Controller 1 Volume Not Ok Fault FB1[260].20'; 8341 '~S001R03CN.I.Slr1PurgeFlt - Seal Controller 1 Purge Fault FB1[260].21'; 8342 '~S001R03CN.I.Slr1DoserNot Filled - Seal Cntrl 1 Doser Not Filled FB1[260].22'; 8343 '~S001R03CN.I.Slr1No2ClnMxr - Seal Cntrl1 No 2C In Mixer Fault FB1[260].23'; 8344 '~S001R03CN.I.Slr1NzlBroken - Seal Controller 1 Nozzle Broken Fault FB1[260].24'; 8345 '~S001R03CN.I.Slr1NozzleChgReq - Seal Cntrl1 Nozzle Change Reqd FB1[260].25'; 8346 '~S001R03CN.I.Slr1CycleInterrupted - Seal Cntrl1 Cycle Interrupted FB1[260].26'; 8347 '~S001R03CN.I.Stdw1Flt - Stud Weld 1 Weld Fault FB1[260].27'; 8348 '~S001R03CN.I.Stdw1DlyExcdd - Stud Weld 1 Time Delay Exceeded Flt FB1[260].28'; 8349 '~S001R03CN.I.Stdw1Maint Reqd - Stud Weld 1 Maintenance Required FB1[260].29'; 8350 '~S001R03CN.I.Stdw1Reject - Stud Weld 1 art Reject Fault FB1[260].30'; 8351 '~S001R03CN.I.Rvt1Flt - Rivet Controller 1 Fault FB1[260].31'; 8352 '~S001R03CN.I.Rvt1DlyExcdd - Rivet Cntrl 1 Time Delay Exceeded Flt FB1[261].0'; 8353 '~S001R03CN.I.AutoPulledTipByp1 - Auto Pulled Tip Bypass 1 FB1[261].1'; 8354 '~S001R03CN.I.StdWld1EquipmentFlt - Stud Weld 1 Equipment Fault FB1[261].2'; 8355 '~S001R03CN.I.StdWld1BrcktNotPresent - Stud Weld 1 Bracket Not Pres FB1[261].3'; 8356 '~S001R03CN.I.PierceFlt - Pierce Fault FB1[261].4'; 8357 '~S001R03CN.I.NoVisionMeasErr - Vision System Measurement Error FB1[261].5'; 8358 '~S001R03CN.I.VisionSysCalErr - Vision System Calibration Fault FB1[261].6'; 8359 '~S001R03CN.I.VisionSysErr - Vision System Error FB1[261].7'; 8360 '~S001R03CN.I.RackOutOfTolerance - Vision Sys Rack Out Of Tolerance FB1[261].8'; 8361 '~S001R03CN.Ix.TorqFlt - Torque Not Ok FB1[261].9'; 8362 '~S001R03CN.Ix.MwFlt - Mig Weld Controller Fault FB1[261].10'; 8363 '~S001R03CN.Ix.MwWireStuckFlt - Mig Welder Wire Stuck FB1[261].11'; 8364 '~S001R03CN.Ix.MwWldFlt - Mig Welder Bad Bronze Weld Indicator Flt FB1[261].12'; 8365 '~S001R03CN.I.O.TipChngReqd1 - Weld Cntrl 1 Tip Change Required FB1[261].13'; 8366 '~S001R03CN.I.M.NutDetectFlt1 - Nut Welder 1 Nut Detection Fault FB1[261].14'; 8367 '~S001R03CN.I.M.NutProjFlt1 - Nut Welder 1 Weld Not In Tolerance FB1[261].15'; 8368 '~S001R03CN.M.WrongRivetAtNose - Remove Wrong Rivet At Nose FB1[261].16'; 8369 '~S001R03CN.Ix.MwWldLimitErr - Mig Welder CurrentVoltage Out of Tolerance FB1[261].17'; 8370 '~S001R03CN.Ix.MigRdy Mig Welder Not Ready FB1[261].18'; 8371 '~Spare FB1[261].19'; 8372 '~Spare FB1[261].20'; 8373 '~S001R03CN.I.Wc2WldFlt -Weld Controller 2 Weld Fault FB1[261].21'; 8374 '~S001R03CN.I.Wc2Flt - Weld Timer Flt - Depress Man Weld To Continue FB1[261].22'; 8375 '~S001R03CN.I.Wc2SGunFlt - Weld Controller 2 Servo Gun Fault FB1[261].23'; 8376 '~S001R03CN.I.Wc2SGunMtrTempFlt - Cntrl 2 Servo Gun Motor Over Temp FB1[261].24'; 8377 '~S001R03CN.I.Td2MtrFlt - Tip Dress 2 Motor Fault FB1[261].25'; 8378 '~S001R03CN.I.WC2XfmrTempFlt - Weld Cntrl 2 Transformer Over Temp FB1[261].26'; 8379 '~S001R03CN.I.AutoTipChng2Flt - Auto Tip Changer 2 Fault FB1[261].27'; 8380 '~S001R03CN.I.Slr2NotReady - Seal Controller 2 Not Ready FB1[261].28'; 8381 '~S001R03CN.I.Slr2MajorFlt - Seal Controller 2 Major Fault FB1[261].29'; 8382 '~S001R03CN.I.Slr2VolNotOk - Seal Controller 2 Volume Not Ok Fault FB1[261].30'; 8383 '~S001R03CN.I.Slr2PurgeFlt - Seal Controller 2 Purge Fault FB1[261].31'; 8384 '~S001R03CN.I.Slr2DoserNot Filled - Seal Cntrl 2 Doser Not Filled FB1[262].0'; 8385 '~S001R03CN.I.Slr2No2ClnMxr - Seal Cntrl2 No 2C In Mixer Fault FB1[262].1'; 8386 '~S001R03CN.I.Slr2NzlBroken - Seal Controller 2 Nozzle Broken Fault FB1[262].2'; 8387 '~S001R03CN.I.Slr2NozzleChgReq - Seal Cntrl2 Nozzle Change Reqd FB1[262].3'; 8388 '~S001R03CN.I.Slr2CycleInterrupted - Seal Cntrl2 Cycle Interrupted FB1[262].4'; 8389 '~S001R03CN.I.Stdw2Flt - Stud Weld 2 Weld Fault FB1[262].5'; 8390 '~S001R03CN.I.Stdw2DlyExcdd - Stud Weld 2 Time Delay Exceeded Flt FB1[262].6'; 8391 '~S001R03CN.I.Stdw2Maint Reqd - Stud Weld 2 Maintenance Required FB1[262].7'; 8392 '~S001R03CN.I.Stdw2Reject - Stud Weld 2 art Reject Fault FB1[262].8'; 8393 '~S001R03CN.I.Rvt2Flt - Rivet Controller 2 Fault FB1[262].9'; 8394 '~S001R03CN.I.Rvt2DlyExcdd - Rivet Cntrl 2 Time Delay Exceeded Flt FB1[262].10'; 8395 '~S001R03CN.I.AutoPulledTipByp2 - Auto Pulled Tip Bypass 2 FB1[262].11'; 8396 '~S001R03CN.I.StdWld2EquipmentFlt - Stud Weld 2 Equipment Fault FB1[262].12'; 8397 '~S001R03CN.I.StdWld2BrcktNotPresent - Stud Weld 2 Bracket Not Pres FB1[262].13'; 8398 '~S001R03CN.Ix.LsrWldMntrFlt - Seam Geometry/Laser Weld Monitor Flt FB1[262].14'; 8399 '~S001R03CN.Ix.LsrHeadFlt - Laser Head Fault FB1[262].15'; 8400 '~S001R03CN.Ix.LsrGlsFlt - Glass Fault FB1[262].16'; 8401 '~S001R03CN.Ix.LsrWhlFlt - Pressure Wheel Not In Range Fault FB1[262].17'; 8402 '~S001R03CN.Ix.LsrGeoFlt - Seam Geometry/Laser Bad Process Geo Flt FB1[262].18'; 8403 '~S001R03CN.Ix.LsrHdCollFlt - Laser Head Collision Fault FB1[262].19'; 8404 '~S001R03CN.Ix.LsrHdSysFlt - Laser Head System Fault FB1[262].20'; 8405 '~S001R03CN.Ix.LsrHdFar - Laser Head Far Fault FB1[262].21'; 8406 '~S001R03CN.Ix.LsrHdSftCollFlt - Laser Head Software Collision Flt FB1[262].22'; 8407 '~S001R03CN.I.O.TipChngReqd2 - Weld Cntrl 2 Tip Change Required FB1[262].23'; 8408 '~S001R03CN.I.M.NutDetectFlt2 - Nut Welder 2 Nut Detection Fault FB1[262].24'; 8409 '~S001R03CN.I.M.NutProjFlt2 - Nut Welder 2 Weld Not In Tolerance FB1[262].25'; 8410 '~S001R03CN.I.TCWrongToolInStand - Tool Changer Wrong Tool In Stand FB1[262].26'; 8411 '~Spare FB1[262].27'; 8412 '~Spare FB1[262].28'; 8413 '~Spare FB1[262].29'; 8414 '~Spare FB1[262].30'; 8415 '~Spare FB1[262].31'; 8416 '~S001R03CN.I.VisionCommOK - Vision System Comm Fault FB1[263].0'; 8417 '~S001R03CN.I.OutOfTolerance - Vision System Out Of Tolerance FB1[263].1'; 8418 '~S001R03CN.I.MeasureReject - Vision System Measure Reject FB1[263].2'; 8419 '~S001R03CN.I.VisionSysCalibrationFlt - Vision System Calibration Flt FB1[263].3'; 8420 '~S001R03CN.I.VisionSysFlt - Vision System Flt FB1[263].4'; 8421 '~Spare FB1[263].5'; 8422 '~Spare FB1[263].6'; 8423 '~Spare FB1[263].7'; 8424 '~Spare FB1[263].8'; 8425 '~Spare FB1[263].9'; 8426 '~Spare FB1[263].10'; 8427 '~Spare FB1[263].11'; 8428 '~Spare FB1[263].12'; 8429 '~Spare FB1[263].13'; 8430 '~Spare FB1[263].14'; 8431 '~Spare FB1[263].15'; 8432 '~Spare FB1[263].16'; 8433 '~Spare FB1[263].17'; 8434 '~S001R03CN.M.InteruptCyc - Laser Cyc Interupt Cut Wire And Reject Car FB1[263].18'; 8435 '~S001R03CN.M.SuspectPart Inspect Vehicle And Accept Or Reject FB1[263].19'; 8436 '~S001R03 Power Meter High Power Fault Detected FB1[263].20'; 8437 '~S001R03 Power Meter Low Power Fault Detected FB1[263].21'; 8438 '~Spare FB1[263].22'; 8439 '~Spare FB1[263].23'; 8440 '~Spare FB1[263].24'; 8441 '~Spare FB1[263].25'; 8442 '~Spare FB1[263].26'; 8443 '~Spare FB1[263].27'; 8444 '~Spare FB1[263].28'; 8445 '~Spare FB1[263].29'; 8446 '~Spare FB1[263].30'; 8447 '~Spare FB1[263].31'; 8448 '~Spare FB1[264].0'; 8449 '~Spare FB1[264].1'; 8450 '~Spare FB1[264].2'; 8451 '~Spare FB1[264].3'; 8452 '~Spare FB1[264].4'; 8453 '~Spare FB1[264].5'; 8454 '~Spare FB1[264].6'; 8455 '~Spare FB1[264].7'; 8456 '~Spare FB1[264].8'; 8457 '~Spare FB1[264].9'; 8458 '~Spare FB1[264].10'; 8459 '~Spare FB1[264].11'; 8460 '~Spare FB1[264].12'; 8461 '~Spare FB1[264].13'; 8462 '~Spare FB1[264].14'; 8463 '~Spare FB1[264].15'; 8464 '~Spare FB1[264].16'; 8465 '~Spare FB1[264].17'; 8466 '~Spare FB1[264].18'; 8467 '~Spare FB1[264].19'; 8468 '~Spare FB1[264].20'; 8469 '~Spare FB1[264].21'; 8470 '~Spare FB1[264].22'; 8471 '~Spare FB1[264].23'; 8472 '~Spare FB1[264].24'; 8473 '~Spare FB1[264].25'; 8474 '~Spare FB1[264].26'; 8475 '~Spare FB1[264].27'; 8476 '~Spare FB1[264].28'; 8477 '~Spare FB1[264].29'; 8478 '~Spare FB1[264].30'; 8479 '~Spare FB1[264].31'; 8480 '~Spare FB1[265].0'; 8481 '~Spare FB1[265].1'; 8482 '~Spare FB1[265].2'; 8483 '~Spare FB1[265].3'; 8484 '~Spare FB1[265].4'; 8485 '~Spare FB1[265].5'; 8486 '~Spare FB1[265].6'; 8487 '~Spare FB1[265].7'; 8488 '~Spare FB1[265].8'; 8489 '~Spare FB1[265].9'; 8490 '~Spare FB1[265].10'; 8491 '~Spare FB1[265].11'; 8492 '~Spare FB1[265].12'; 8493 '~Spare FB1[265].13'; 8494 '~Spare FB1[265].14'; 8495 '~Spare FB1[265].15'; 8496 '~Spare FB1[265].16'; 8497 '~Spare FB1[265].17'; 8498 '~Spare FB1[265].18'; 8499 '~Spare FB1[265].19'; 8500 '~Spare FB1[265].20'; 8501 '~Spare FB1[265].21'; 8502 '~Spare FB1[265].22'; 8503 '~Spare FB1[265].23'; 8504 '~Spare FB1[265].24'; 8505 '~Spare FB1[265].25'; 8506 '~Spare FB1[265].26'; 8507 '~Spare FB1[265].27'; 8508 '~Spare FB1[265].28'; 8509 '~Spare FB1[265].29'; 8510 '~Spare FB1[265].30'; 8511 '~Spare FB1[265].31'; 8512 '~Spare FB1[266].0'; 8513 '~Spare FB1[266].1'; 8514 '~Spare FB1[266].2'; 8515 '~Spare FB1[266].3'; 8516 '~Spare FB1[266].4'; 8517 '~Spare FB1[266].5'; 8518 '~Spare FB1[266].6'; 8519 '~Spare FB1[266].7'; 8520 '~Spare FB1[266].8'; 8521 '~Spare FB1[266].9'; 8522 '~Spare FB1[266].10'; 8523 '~Spare FB1[266].11'; 8524 '~Spare FB1[266].12'; 8525 '~Spare FB1[266].13'; 8526 '~Spare FB1[266].14'; 8527 '~Spare FB1[266].15'; 8528 '~Spare FB1[266].16'; 8529 '~Spare FB1[266].17'; 8530 '~Spare FB1[266].18'; 8531 '~Spare FB1[266].19'; 8532 '~Spare FB1[266].20'; 8533 '~Spare FB1[266].21'; 8534 '~Spare FB1[266].22'; 8535 '~Spare FB1[266].23'; 8536 '~Spare FB1[266].24'; 8537 '~Spare FB1[266].25'; 8538 '~Spare FB1[266].26'; 8539 '~Spare FB1[266].27'; 8540 '~Spare FB1[266].28'; 8541 '~Spare FB1[266].29'; 8542 '~Spare FB1[266].30'; 8543 '~Spare FB1[266].31'; 8544 '~Spare FB1[267].0'; 8545 '~Spare FB1[267].1'; 8546 '~Spare FB1[267].2'; 8547 '~Spare FB1[267].3'; 8548 '~Spare FB1[267].4'; 8549 '~Spare FB1[267].5'; 8550 '~Spare FB1[267].6'; 8551 '~Spare FB1[267].7'; 8552 '~Spare FB1[267].8'; 8553 '~Spare FB1[267].9'; 8554 '~Spare FB1[267].10'; 8555 '~Spare FB1[267].11'; 8556 '~Spare FB1[267].12'; 8557 '~Spare FB1[267].13'; 8558 '~Spare FB1[267].14'; 8559 '~Spare FB1[267].15'; 8560 '~Spare FB1[267].16'; 8561 '~Spare FB1[267].17'; 8562 '~Spare FB1[267].18'; 8563 '~Spare FB1[267].19'; 8564 '~Spare FB1[267].20'; 8565 '~Spare FB1[267].21'; 8566 '~Spare FB1[267].22'; 8567 '~Spare FB1[267].23'; 8568 '~Spare FB1[267].24'; 8569 '~Spare FB1[267].25'; 8570 '~Spare FB1[267].26'; 8571 '~Spare FB1[267].27'; 8572 '~Spare FB1[267].28'; 8573 '~Spare FB1[267].29'; 8574 '~Spare FB1[267].30'; 8575 '~Spare FB1[267].31'; 8576 '~S001R04CN.I.RbtCtrlFlt - Control Fault FB1[268].0'; 8577 '~S001R04CN.I.CollDetect - Collision Detect FB1[268].1'; 8578 '~S001R04CN.Ix.RbtPromptBox - View Prompt Box at Teach Pendant FB1[268].2'; 8579 '~Spare FB1[268].3'; 8580 '~Spare FB1[268].4'; 8581 '~Spare FB1[268].5'; 8582 '~Spare FB1[268].6'; 8583 '~Spare FB1[268].7'; 8584 '~Spare FB1[268].8'; 8585 '~Spare FB1[268].9'; 8586 '~Spare FB1[268].10'; 8587 '~S001R04CN.I.Wc1WldFlt -Weld Controller 1 Weld Fault FB1[268].11'; 8588 '~S001R04CN.I.Wc1Flt - Weld Timer Flt - Depress Man Weld To Continue FB1[268].12'; 8589 '~S001R04CN.I.Wc1SGunFlt - Weld Controller 1 Servo Gun Fault FB1[268].13'; 8590 '~S001R04CN.I.Wc1SGunMtrTempFlt - Cntrl 1 Servo Gun Motor Over Temp FB1[268].14'; 8591 '~S001R04CN.I.Td1MtrFlt - Tip Dress 1 Motor Fault FB1[268].15'; 8592 '~S001R04CN.I.WC1XfmrTempFlt - Weld Cntrl 1 Transformer Over Temp FB1[268].16'; 8593 '~S001R04CN.I.AutoTipChng1Flt - Auto Tip Changer 1 Fault FB1[268].17'; 8594 '~S001R04CN.I.Slr1NotReady - Seal Controller 1 Not Ready FB1[268].18'; 8595 '~S001R04CN.I.Slr1MajorFlt - Seal Controller 1 Major Fault FB1[268].19'; 8596 '~S001R04CN.I.Slr1VolNotOk - Seal Controller 1 Volume Not Ok Fault FB1[268].20'; 8597 '~S001R04CN.I.Slr1PurgeFlt - Seal Controller 1 Purge Fault FB1[268].21'; 8598 '~S001R04CN.I.Slr1DoserNot Filled - Seal Cntrl 1 Doser Not Filled FB1[268].22'; 8599 '~S001R04CN.I.Slr1No2ClnMxr - Seal Cntrl1 No 2C In Mixer Fault FB1[268].23'; 8600 '~S001R04CN.I.Slr1NzlBroken - Seal Controller 1 Nozzle Broken Fault FB1[268].24'; 8601 '~S001R04CN.I.Slr1NozzleChgReq - Seal Cntrl1 Nozzle Change Reqd FB1[268].25'; 8602 '~S001R04CN.I.Slr1CycleInterrupted - Seal Cntrl1 Cycle Interrupted FB1[268].26'; 8603 '~S001R04CN.I.Stdw1Flt - Stud Weld 1 Weld Fault FB1[268].27'; 8604 '~S001R04CN.I.Stdw1DlyExcdd - Stud Weld 1 Time Delay Exceeded Flt FB1[268].28'; 8605 '~S001R04CN.I.Stdw1Maint Reqd - Stud Weld 1 Maintenance Required FB1[268].29'; 8606 '~S001R04CN.I.Stdw1Reject - Stud Weld 1 art Reject Fault FB1[268].30'; 8607 '~S001R04CN.I.Rvt1Flt - Rivet Controller 1 Fault FB1[268].31'; 8608 '~S001R04CN.I.Rvt1DlyExcdd - Rivet Cntrl 1 Time Delay Exceeded Flt FB1[269].0'; 8609 '~S001R04CN.I.AutoPulledTipByp1 - Auto Pulled Tip Bypass 1 FB1[269].1'; 8610 '~S001R04CN.I.StdWld1EquipmentFlt - Stud Weld 1 Equipment Fault FB1[269].2'; 8611 '~S001R04CN.I.StdWld1BrcktNotPresent - Stud Weld 1 Bracket Not Pres FB1[269].3'; 8612 '~S001R04CN.I.PierceFlt - Pierce Fault FB1[269].4'; 8613 '~S001R04CN.I.NoVisionMeasErr - Vision System Measurement Error FB1[269].5'; 8614 '~S001R04CN.I.VisionSysCalErr - Vision System Calibration Fault FB1[269].6'; 8615 '~S001R04CN.I.VisionSysErr - Vision System Error FB1[269].7'; 8616 '~S001R04CN.I.RackOutOfTolerance - Vision Sys Rack Out Of Tolerance FB1[269].8'; 8617 '~S001R04CN.Ix.TorqFlt - Torque Not Ok FB1[269].9'; 8618 '~S001R04CN.Ix.MwFlt - Mig Weld Controller Fault FB1[269].10'; 8619 '~S001R04CN.Ix.MwWireStuckFlt - Mig Welder Wire Stuck FB1[269].11'; 8620 '~S001R04CN.Ix.MwWldFlt - Mig Welder Bad Bronze Weld Indicator Flt FB1[269].12'; 8621 '~S001R04CN.I.O.TipChngReqd1 - Weld Cntrl 1 Tip Change Required FB1[269].13'; 8622 '~S001R04CN.I.M.NutDetectFlt1 - Nut Welder 1 Nut Detection Fault FB1[269].14'; 8623 '~S001R04CN.I.M.NutProjFlt1 - Nut Welder 1 Weld Not In Tolerance FB1[269].15'; 8624 '~S001R04CN.M.WrongRivetAtNose - Remove Wrong Rivet At Nose FB1[269].16'; 8625 '~S001R04CN.Ix.MwWldLimitErr - Mig Welder CurrentVoltage Out of Tolerance FB1[269].17'; 8626 '~S001R04CN.Ix.MigRdy Mig Welder Not Ready FB1[269].18'; 8627 '~Spare FB1[269].19'; 8628 '~Spare FB1[269].20'; 8629 '~S001R04CN.I.Wc2WldFlt -Weld Controller 2 Weld Fault FB1[269].21'; 8630 '~S001R04CN.I.Wc2Flt - Weld Timer Flt - Depress Man Weld To Continue FB1[269].22'; 8631 '~S001R04CN.I.Wc2SGunFlt - Weld Controller 2 Servo Gun Fault FB1[269].23'; 8632 '~S001R04CN.I.Wc2SGunMtrTempFlt - Cntrl 2 Servo Gun Motor Over Temp FB1[269].24'; 8633 '~S001R04CN.I.Td2MtrFlt - Tip Dress 2 Motor Fault FB1[269].25'; 8634 '~S001R04CN.I.WC2XfmrTempFlt - Weld Cntrl 2 Transformer Over Temp FB1[269].26'; 8635 '~S001R04CN.I.AutoTipChng2Flt - Auto Tip Changer 2 Fault FB1[269].27'; 8636 '~S001R04CN.I.Slr2NotReady - Seal Controller 2 Not Ready FB1[269].28'; 8637 '~S001R04CN.I.Slr2MajorFlt - Seal Controller 2 Major Fault FB1[269].29'; 8638 '~S001R04CN.I.Slr2VolNotOk - Seal Controller 2 Volume Not Ok Fault FB1[269].30'; 8639 '~S001R04CN.I.Slr2PurgeFlt - Seal Controller 2 Purge Fault FB1[269].31'; 8640 '~S001R04CN.I.Slr2DoserNot Filled - Seal Cntrl 2 Doser Not Filled FB1[270].0'; 8641 '~S001R04CN.I.Slr2No2ClnMxr - Seal Cntrl2 No 2C In Mixer Fault FB1[270].1'; 8642 '~S001R04CN.I.Slr2NzlBroken - Seal Controller 2 Nozzle Broken Fault FB1[270].2'; 8643 '~S001R04CN.I.Slr2NozzleChgReq - Seal Cntrl2 Nozzle Change Reqd FB1[270].3'; 8644 '~S001R04CN.I.Slr2CycleInterrupted - Seal Cntrl2 Cycle Interrupted FB1[270].4'; 8645 '~S001R04CN.I.Stdw2Flt - Stud Weld 2 Weld Fault FB1[270].5'; 8646 '~S001R04CN.I.Stdw2DlyExcdd - Stud Weld 2 Time Delay Exceeded Flt FB1[270].6'; 8647 '~S001R04CN.I.Stdw2Maint Reqd - Stud Weld 2 Maintenance Required FB1[270].7'; 8648 '~S001R04CN.I.Stdw2Reject - Stud Weld 2 art Reject Fault FB1[270].8'; 8649 '~S001R04CN.I.Rvt2Flt - Rivet Controller 2 Fault FB1[270].9'; 8650 '~S001R04CN.I.Rvt2DlyExcdd - Rivet Cntrl 2 Time Delay Exceeded Flt FB1[270].10'; 8651 '~S001R04CN.I.AutoPulledTipByp2 - Auto Pulled Tip Bypass 2 FB1[270].11'; 8652 '~S001R04CN.I.StdWld2EquipmentFlt - Stud Weld 2 Equipment Fault FB1[270].12'; 8653 '~S001R04CN.I.StdWld2BrcktNotPresent - Stud Weld 2 Bracket Not Pres FB1[270].13'; 8654 '~S001R04CN.Ix.LsrWldMntrFlt - Seam Geometry/Laser Weld Monitor Flt FB1[270].14'; 8655 '~S001R04CN.Ix.LsrHeadFlt - Laser Head Fault FB1[270].15'; 8656 '~S001R04CN.Ix.LsrGlsFlt - Glass Fault FB1[270].16'; 8657 '~S001R04CN.Ix.LsrWhlFlt - Pressure Wheel Not In Range Fault FB1[270].17'; 8658 '~S001R04CN.Ix.LsrGeoFlt - Seam Geometry/Laser Bad Process Geo Flt FB1[270].18'; 8659 '~S001R04CN.Ix.LsrHdCollFlt - Laser Head Collision Fault FB1[270].19'; 8660 '~S001R04CN.Ix.LsrHdSysFlt - Laser Head System Fault FB1[270].20'; 8661 '~S001R04CN.Ix.LsrHdFar - Laser Head Far Fault FB1[270].21'; 8662 '~S001R04CN.Ix.LsrHdSftCollFlt - Laser Head Software Collision Flt FB1[270].22'; 8663 '~S001R04CN.I.O.TipChngReqd2 - Weld Cntrl 2 Tip Change Required FB1[270].23'; 8664 '~S001R04CN.I.M.NutDetectFlt2 - Nut Welder 2 Nut Detection Fault FB1[270].24'; 8665 '~S001R04CN.I.M.NutProjFlt2 - Nut Welder 2 Weld Not In Tolerance FB1[270].25'; 8666 '~S001R04CN.I.TCWrongToolInStand - Tool Changer Wrong Tool In Stand FB1[270].26'; 8667 '~Spare FB1[270].27'; 8668 '~Spare FB1[270].28'; 8669 '~Spare FB1[270].29'; 8670 '~Spare FB1[270].30'; 8671 '~Spare FB1[270].31'; 8672 '~S001R04CN.I.VisionCommOK - Vision System Comm Fault FB1[271].0'; 8673 '~S001R04CN.I.OutOfTolerance - Vision System Out Of Tolerance FB1[271].1'; 8674 '~S001R04CN.I.MeasureReject - Vision System Measure Reject FB1[271].2'; 8675 '~S001R04CN.I.VisionSysCalibrationFlt - Vision System Calibration Flt FB1[271].3'; 8676 '~S001R04CN.I.VisionSysFlt - Vision System Flt FB1[271].4'; 8677 '~Spare FB1[271].5'; 8678 '~Spare FB1[271].6'; 8679 '~Spare FB1[271].7'; 8680 '~Spare FB1[271].8'; 8681 '~Spare FB1[271].9'; 8682 '~Spare FB1[271].10'; 8683 '~Spare FB1[271].11'; 8684 '~Spare FB1[271].12'; 8685 '~Spare FB1[271].13'; 8686 '~Spare FB1[271].14'; 8687 '~Spare FB1[271].15'; 8688 '~Spare FB1[271].16'; 8689 '~Spare FB1[271].17'; 8690 '~S001R04CN.M.InteruptCyc - Laser Cyc Interupt Cut Wire And Reject Car FB1[271].18'; 8691 '~S001R04CN.M.SuspectPart Inspect Vehicle And Accept Or Reject FB1[271].19'; 8692 '~S001R04 Power Meter High Power Fault Detected FB1[271].20'; 8693 '~S001R04 Power Meter Low Power Fault Detected FB1[271].21'; 8694 '~Spare FB1[271].22'; 8695 '~Spare FB1[271].23'; 8696 '~Spare FB1[271].24'; 8697 '~Spare FB1[271].25'; 8698 '~Spare FB1[271].26'; 8699 '~Spare FB1[271].27'; 8700 '~Spare FB1[271].28'; 8701 '~Spare FB1[271].29'; 8702 '~Spare FB1[271].30'; 8703 '~Spare FB1[271].31'; 8704 '~Spare FB1[272].0'; 8705 '~Spare FB1[272].1'; 8706 '~Spare FB1[272].2'; 8707 '~Spare FB1[272].3'; 8708 '~Spare FB1[272].4'; 8709 '~Spare FB1[272].5'; 8710 '~Spare FB1[272].6'; 8711 '~Spare FB1[272].7'; 8712 '~Spare FB1[272].8'; 8713 '~Spare FB1[272].9'; 8714 '~Spare FB1[272].10'; 8715 '~Spare FB1[272].11'; 8716 '~Spare FB1[272].12'; 8717 '~Spare FB1[272].13'; 8718 '~Spare FB1[272].14'; 8719 '~Spare FB1[272].15'; 8720 '~Spare FB1[272].16'; 8721 '~Spare FB1[272].17'; 8722 '~Spare FB1[272].18'; 8723 '~Spare FB1[272].19'; 8724 '~Spare FB1[272].20'; 8725 '~Spare FB1[272].21'; 8726 '~Spare FB1[272].22'; 8727 '~Spare FB1[272].23'; 8728 '~Spare FB1[272].24'; 8729 '~Spare FB1[272].25'; 8730 '~Spare FB1[272].26'; 8731 '~Spare FB1[272].27'; 8732 '~Spare FB1[272].28'; 8733 '~Spare FB1[272].29'; 8734 '~Spare FB1[272].30'; 8735 '~Spare FB1[272].31'; 8736 '~Spare FB1[273].0'; 8737 '~Spare FB1[273].1'; 8738 '~Spare FB1[273].2'; 8739 '~Spare FB1[273].3'; 8740 '~Spare FB1[273].4'; 8741 '~Spare FB1[273].5'; 8742 '~Spare FB1[273].6'; 8743 '~Spare FB1[273].7'; 8744 '~Spare FB1[273].8'; 8745 '~Spare FB1[273].9'; 8746 '~Spare FB1[273].10'; 8747 '~Spare FB1[273].11'; 8748 '~Spare FB1[273].12'; 8749 '~Spare FB1[273].13'; 8750 '~Spare FB1[273].14'; 8751 '~Spare FB1[273].15'; 8752 '~Spare FB1[273].16'; 8753 '~Spare FB1[273].17'; 8754 '~Spare FB1[273].18'; 8755 '~Spare FB1[273].19'; 8756 '~Spare FB1[273].20'; 8757 '~Spare FB1[273].21'; 8758 '~Spare FB1[273].22'; 8759 '~Spare FB1[273].23'; 8760 '~Spare FB1[273].24'; 8761 '~Spare FB1[273].25'; 8762 '~Spare FB1[273].26'; 8763 '~Spare FB1[273].27'; 8764 